(* Logix 5000 project; controller MV vendor 1 type 14 code 217 rev 31.11; software revision 31.00; part 35 of 53 *)
(* tags used below, declared in another part *)
   Alarm_Reset : BOOL;
   Analog_Fault_No : DINT;
   Analog_Simulation_Enabled : BOOL;
   CWD : CHECKWORD_FLAGS;
   Default_Check_Time : DINT;
   MV_MV18_RTD1_AI : PlantItem;   // MV18_RTD1
   MV_MV18_RTD1_AI_RawInput : ALIAS FOR Remote_IO:3:I.Ch5Data;   // Real Analog Input , Do Not Use In Code
   MV_MV19_RTD1_AI : PlantItem;   // MV19_RTD1
   MV_MV19_RTD1_AI_RawInput : ALIAS FOR Remote_IO:4:I.Ch0Data;   // Real Analog Input , Do Not Use In Code
   MV_MV20_RTD1_AI : PlantItem;   // MV20_RTD1
   MV_MV20_RTD1_AI_RawInput : ALIAS FOR Remote_IO:5:I.Ch1Data;   // Real Analog Input , Do Not Use In Code
   MV_MV21_RTD1_AI : PlantItem;   // MV21_RTD1
   MV_MV21_RTD1_AI_RawInput : ALIAS FOR Remote_IO:5:I.Ch2Data;   // Real Analog Input , Do Not Use In Code
   MV_MV22_RTD1_AI : PlantItem;   // MV22_RTD1
   MV_MV22_RTD1_AI_RawInput : ALIAS FOR Remote_IO:5:I.Ch3Data;   // Real Analog Input , Do Not Use In Code
   MV_MV23_RTD1_AI : PlantItem;   // MV23_RTD1
   MV_MV23_RTD1_AI_RawInput : ALIAS FOR Remote_IO:5:I.Ch4Data;   // Real Analog Input , Do Not Use In Code
   MV_MV30_RTD1_AI : PlantItem;   // MV30_RTD1
   MV_MV30_RTD1_AI_RawInput : ALIAS FOR Remote_IO:4:I.Ch1Data;   // Real Analog Input , Do Not Use In Code
   MV_MV31_RTD1_AI : PlantItem;   // MV31_RTD1
   MV_MV31_RTD1_AI_RawInput : ALIAS FOR Remote_IO:4:I.Ch2Data;   // Real Analog Input , Do Not Use In Code
   MV_MV32_RTD1_AI : PlantItem;   // MV32_RTD1
   MV_MV32_RTD1_AI_RawInput : ALIAS FOR Remote_IO:4:I.Ch3Data;   // Real Analog Input , Do Not Use In Code
   MV_MV33_RTD1_AI : PlantItem;   // MV33_RTD1
   MV_MV33_RTD1_AI_RawInput : ALIAS FOR Remote_IO:4:I.Ch4Data;   // Real Analog Input , Do Not Use In Code
   MV_MV34_RTD1_AI : PlantItem;   // MV34_RTD1
   MV_MV34_RTD1_AI_RawInput : ALIAS FOR Remote_IO:4:I.Ch5Data;   // Real Analog Input , Do Not Use In Code
   MV_MV35_RTD1_AI : PlantItem;   // MV35_RTD1
   MV_MV35_RTD1_AI_RawInput : ALIAS FOR Remote_IO:5:I.Ch0Data;   // Real Analog Input , Do Not Use In Code
   MV_MV36_TTX01_AI : PlantItem;   // MV36_TTX01
   MV_MV36_TTX01_AI_RawInput : ALIAS FOR Remote_IO:7:I.Ch00Data;   // Real Analog Input , Do Not Use In Code
   MV_MV37_TTX01_AI : PlantItem;   // MV37_TTX01
   MV_MV37_TTX01_AI_RawInput : ALIAS FOR Remote_IO:7:I.Ch01Data;   // Real Analog Input , Do Not Use In Code
   MV_MV38_TTX01_AI : PlantItem;   // MV38_TTX01
   MV_MV38_TTX01_AI_RawInput : ALIAS FOR Remote_IO:7:I.Ch02Data;   // Real Analog Input , Do Not Use In Code
   MV_MV39_TTX01_AI : PlantItem;   // MV39_TTX01
   MV_MV39_TTX01_AI_RawInput : ALIAS FOR Remote_IO:7:I.Ch03Data;   // Real Analog Input , Do Not Use In Code
   MV_MV40_TTX01_AI : PlantItem;   // MV40_TTX01
   MV_MV40_TTX01_AI_RawInput : ALIAS FOR Remote_IO:7:I.Ch04Data;   // Real Analog Input , Do Not Use In Code
   MV_MV41_TTX01_AI : PlantItem;   // MV41_TTX01
   MV_MV41_TTX01_AI_RawInput : ALIAS FOR Remote_IO:7:I.Ch05Data;   // Real Analog Input , Do Not Use In Code
   MV_MV42_TTX01_AI : PlantItem;   // MV42_TTX01
   MV_MV42_TTX01_AI_RawInput : ALIAS FOR Remote_IO:7:I.Ch06Data;   // Real Analog Input , Do Not Use In Code
   MV_MV43_TTX01_AI : PlantItem;   // MV43_TTX01
   MV_MV43_TTX01_AI_RawInput : ALIAS FOR Remote_IO:7:I.Ch07Data;   // Real Analog Input , Do Not Use In Code
   MV_MV44_TTX01_AI : PlantItem;   // MV44_TTX01
   MV_MV44_TTX01_AI_RawInput : ALIAS FOR Remote_IO:7:I.Ch08Data;   // Real Analog Input , Do Not Use In Code
   MV_MV45_TTX01_AI : PlantItem;   // MV45_TTX01
   MV_MV45_TTX01_AI_RawInput : ALIAS FOR Remote_IO:7:I.Ch09Data;   // Real Analog Input , Do Not Use In Code
   MV_MV46_TTX01_AI : PlantItem;   // MV46_TTX01
   MV_MV46_TTX01_AI_RawInput : ALIAS FOR Remote_IO:7:I.Ch10Data;   // Real Analog Input , Do Not Use In Code
   MV_MV47_TTX01_AI : PlantItem;   // MV47_TTX01
   MV_MV47_TTX01_AI_RawInput : ALIAS FOR Remote_IO:7:I.Ch11Data;   // Real Analog Input , Do Not Use In Code
   One_Second_One_Scan : ALIAS FOR One_Second_1_scan;
   overrange_RIO_analog_value : REAL;
   underrange_RIO_analog_value : REAL;
(* MV_Common, continued *)

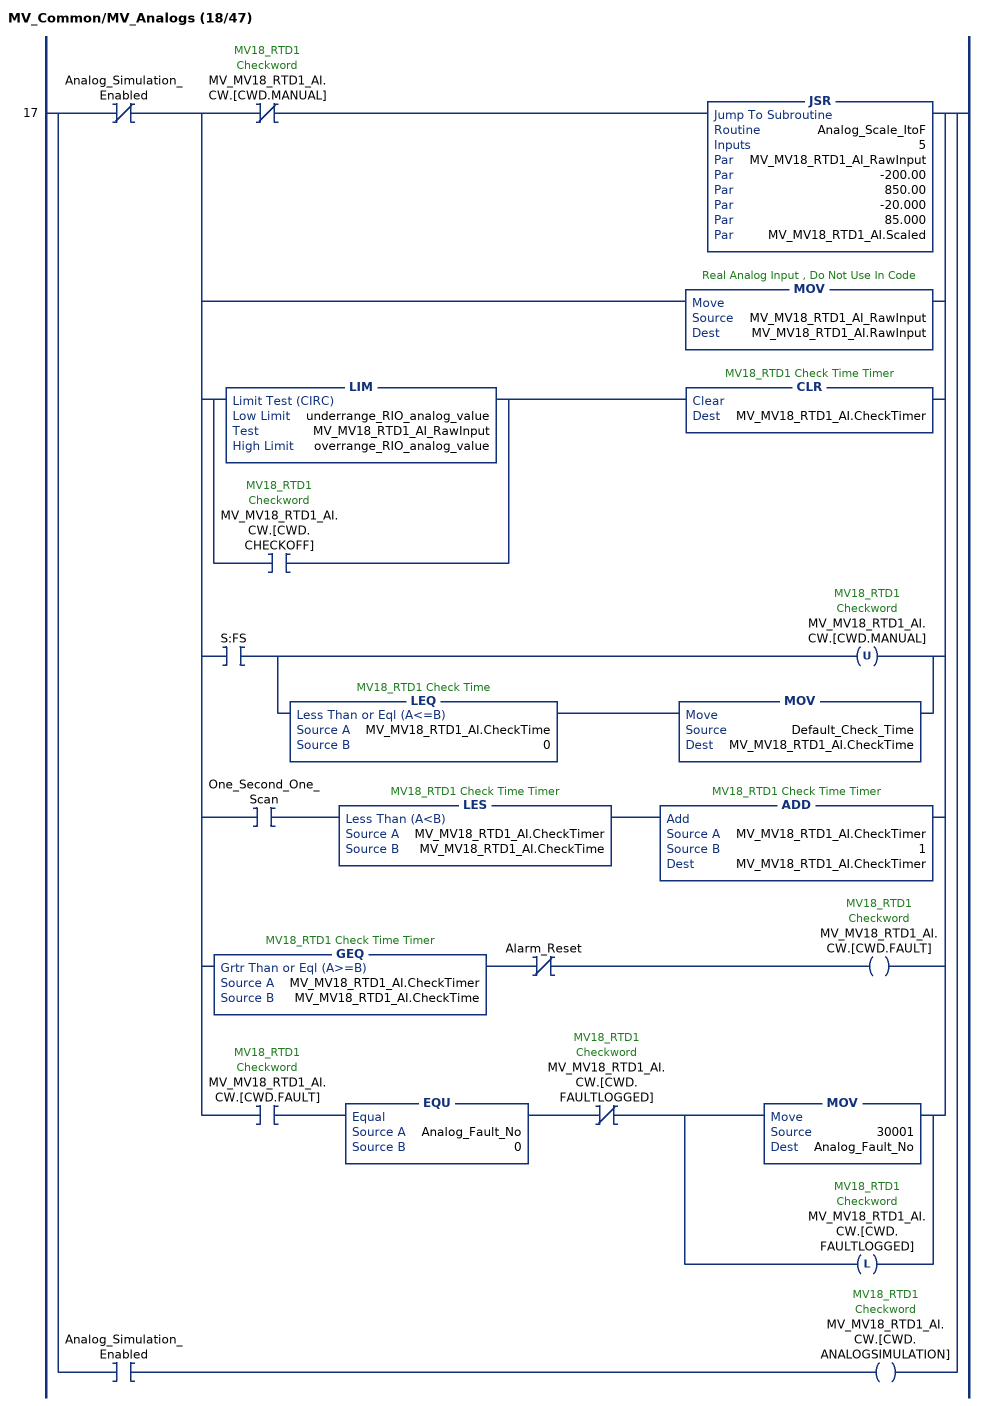
   [picture p810: MV_Common/MV_Analogs rungs 17-17]
   17: [XIO(Analog_Simulation_Enabled) [XIO(MV_MV18_RTD1_AI.CW.[CWD.MANUAL]) JSR(Analog_Scale_ItoF,5,MV_MV18_RTD1_AI_RawInput,-200.00,850.00,-20.000,85.000,MV_MV18_RTD1_AI.Scaled) ,MOV(MV_MV18_RTD1_AI_RawInput,MV_MV18_RTD1_AI.RawInput) ,[LIM(underrange_RIO_analog_value,MV_MV18_RTD1_AI_RawInput,overrange_RIO_analog_value) ,XIC(MV_MV18_RTD1_AI.CW.[CWD.CHECKOFF]) ] CLR(MV_MV18_RTD1_AI.CheckTimer) ,XIC(S:FS) [OTU(MV_MV18_RTD1_AI.CW.[CWD.MANUAL]) ,LEQ(MV_MV18_RTD1_AI.CheckTime,0) MOV(Default_Check_Time,MV_MV18_RTD1_AI.CheckTime) ] ,XIC(One_Second_One_Scan) LES(MV_MV18_RTD1_AI.CheckTimer,MV_MV18_RTD1_AI.CheckTime) ADD(MV_MV18_RTD1_AI.CheckTimer,1,MV_MV18_RTD1_AI.CheckTimer) ,GEQ(MV_MV18_RTD1_AI.CheckTimer,MV_MV18_RTD1_AI.CheckTime) XIO(Alarm_Reset) OTE(MV_MV18_RTD1_AI.CW.[CWD.FAULT]) ,XIC(MV_MV18_RTD1_AI.CW.[CWD.FAULT]) EQU(Analog_Fault_No,0) XIO(MV_MV18_RTD1_AI.CW.[CWD.FAULTLOGGED]) [MOV(30001,Analog_Fault_No) ,OTL(MV_MV18_RTD1_AI.CW.[CWD.FAULTLOGGED]) ] ] ,XIC(Analog_Simulation_Enabled) OTE(MV_MV18_RTD1_AI.CW.[CWD.ANALOGSIMULATION]) ];
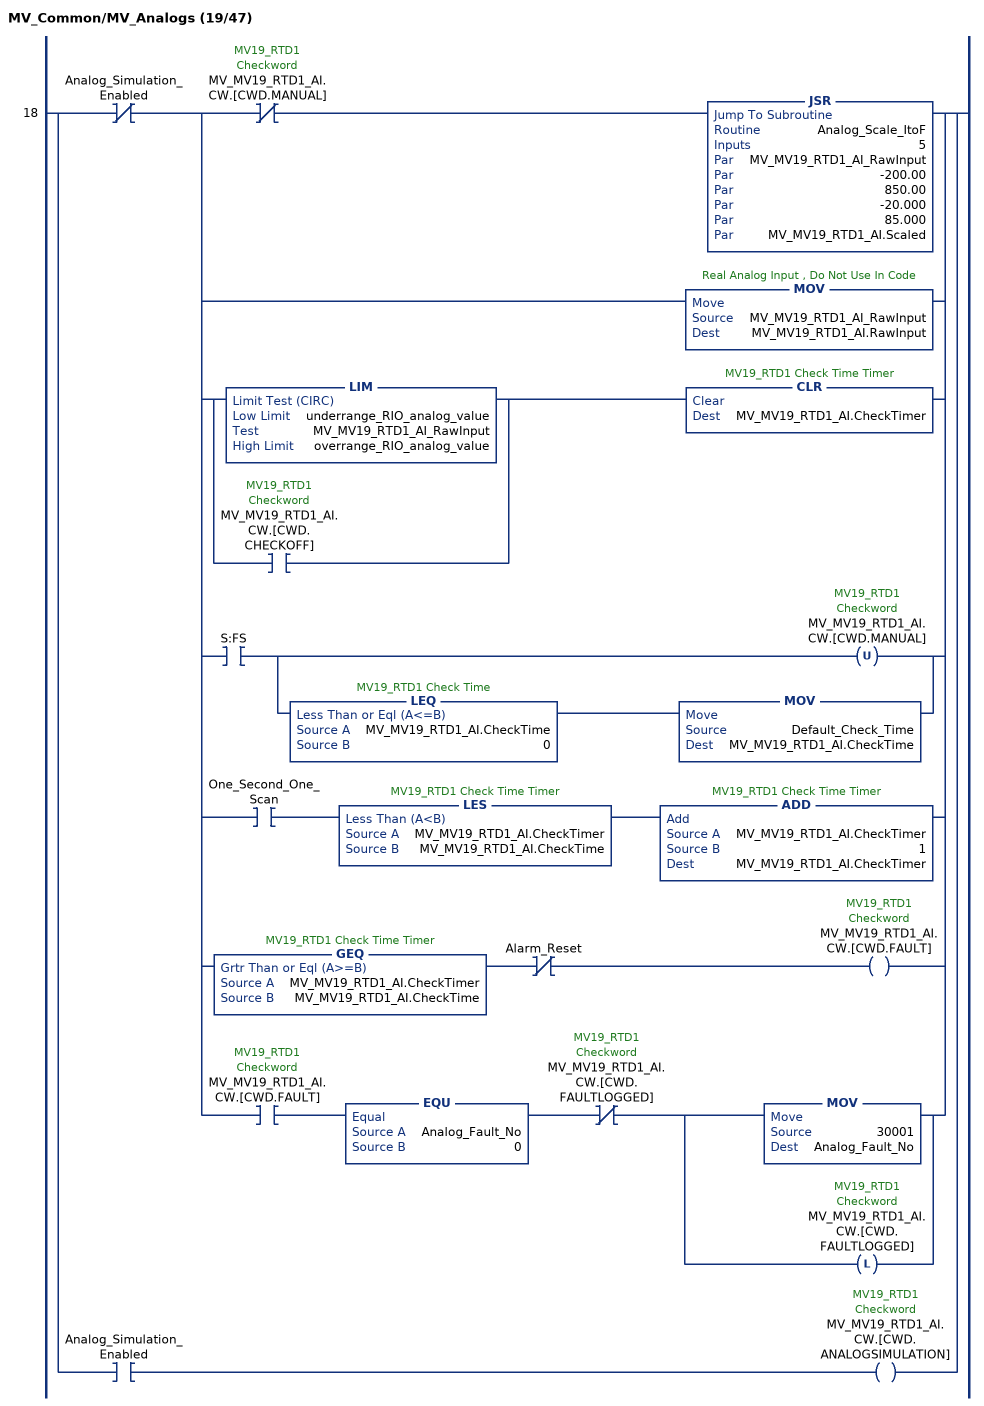
   18: [XIO(Analog_Simulation_Enabled) [XIO(MV_MV19_RTD1_AI.CW.[CWD.MANUAL]) JSR(Analog_Scale_ItoF,5,MV_MV19_RTD1_AI_RawInput,-200.00,850.00,-20.000,85.000,MV_MV19_RTD1_AI.Scaled) ,MOV(MV_MV19_RTD1_AI_RawInput,MV_MV19_RTD1_AI.RawInput) ,[LIM(underrange_RIO_analog_value,MV_MV19_RTD1_AI_RawInput,overrange_RIO_analog_value) ,XIC(MV_MV19_RTD1_AI.CW.[CWD.CHECKOFF]) ] CLR(MV_MV19_RTD1_AI.CheckTimer) ,XIC(S:FS) [OTU(MV_MV19_RTD1_AI.CW.[CWD.MANUAL]) ,LEQ(MV_MV19_RTD1_AI.CheckTime,0) MOV(Default_Check_Time,MV_MV19_RTD1_AI.CheckTime) ] ,XIC(One_Second_One_Scan) LES(MV_MV19_RTD1_AI.CheckTimer,MV_MV19_RTD1_AI.CheckTime) ADD(MV_MV19_RTD1_AI.CheckTimer,1,MV_MV19_RTD1_AI.CheckTimer) ,GEQ(MV_MV19_RTD1_AI.CheckTimer,MV_MV19_RTD1_AI.CheckTime) XIO(Alarm_Reset) OTE(MV_MV19_RTD1_AI.CW.[CWD.FAULT]) ,XIC(MV_MV19_RTD1_AI.CW.[CWD.FAULT]) EQU(Analog_Fault_No,0) XIO(MV_MV19_RTD1_AI.CW.[CWD.FAULTLOGGED]) [MOV(30001,Analog_Fault_No) ,OTL(MV_MV19_RTD1_AI.CW.[CWD.FAULTLOGGED]) ] ] ,XIC(Analog_Simulation_Enabled) OTE(MV_MV19_RTD1_AI.CW.[CWD.ANALOGSIMULATION]) ];
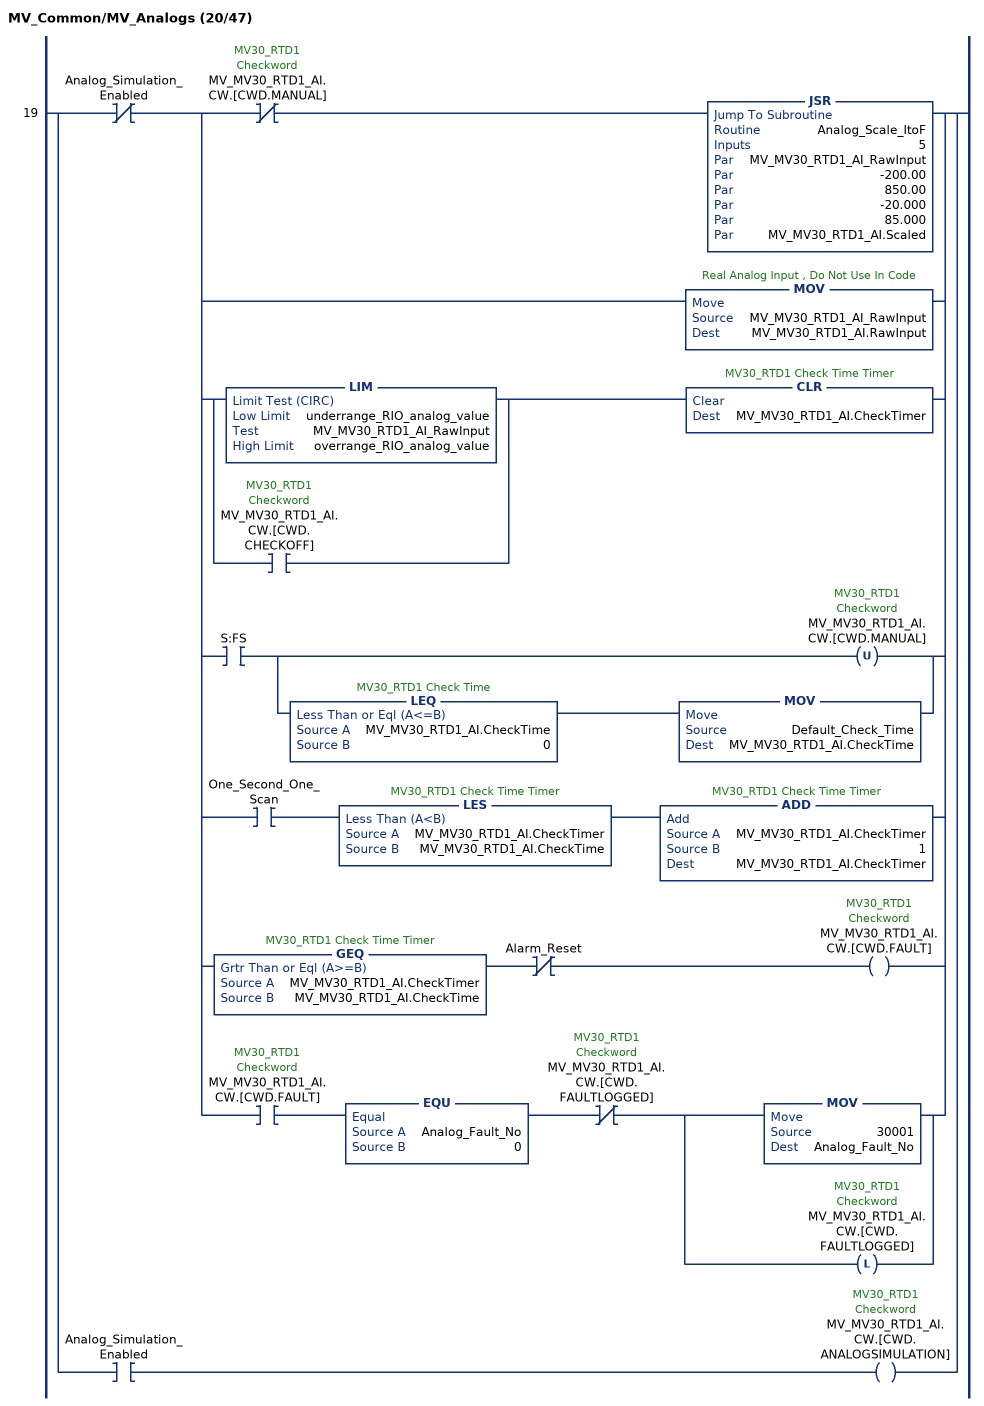
   19: [XIO(Analog_Simulation_Enabled) [XIO(MV_MV30_RTD1_AI.CW.[CWD.MANUAL]) JSR(Analog_Scale_ItoF,5,MV_MV30_RTD1_AI_RawInput,-200.00,850.00,-20.000,85.000,MV_MV30_RTD1_AI.Scaled) ,MOV(MV_MV30_RTD1_AI_RawInput,MV_MV30_RTD1_AI.RawInput) ,[LIM(underrange_RIO_analog_value,MV_MV30_RTD1_AI_RawInput,overrange_RIO_analog_value) ,XIC(MV_MV30_RTD1_AI.CW.[CWD.CHECKOFF]) ] CLR(MV_MV30_RTD1_AI.CheckTimer) ,XIC(S:FS) [OTU(MV_MV30_RTD1_AI.CW.[CWD.MANUAL]) ,LEQ(MV_MV30_RTD1_AI.CheckTime,0) MOV(Default_Check_Time,MV_MV30_RTD1_AI.CheckTime) ] ,XIC(One_Second_One_Scan) LES(MV_MV30_RTD1_AI.CheckTimer,MV_MV30_RTD1_AI.CheckTime) ADD(MV_MV30_RTD1_AI.CheckTimer,1,MV_MV30_RTD1_AI.CheckTimer) ,GEQ(MV_MV30_RTD1_AI.CheckTimer,MV_MV30_RTD1_AI.CheckTime) XIO(Alarm_Reset) OTE(MV_MV30_RTD1_AI.CW.[CWD.FAULT]) ,XIC(MV_MV30_RTD1_AI.CW.[CWD.FAULT]) EQU(Analog_Fault_No,0) XIO(MV_MV30_RTD1_AI.CW.[CWD.FAULTLOGGED]) [MOV(30001,Analog_Fault_No) ,OTL(MV_MV30_RTD1_AI.CW.[CWD.FAULTLOGGED]) ] ] ,XIC(Analog_Simulation_Enabled) OTE(MV_MV30_RTD1_AI.CW.[CWD.ANALOGSIMULATION]) ];
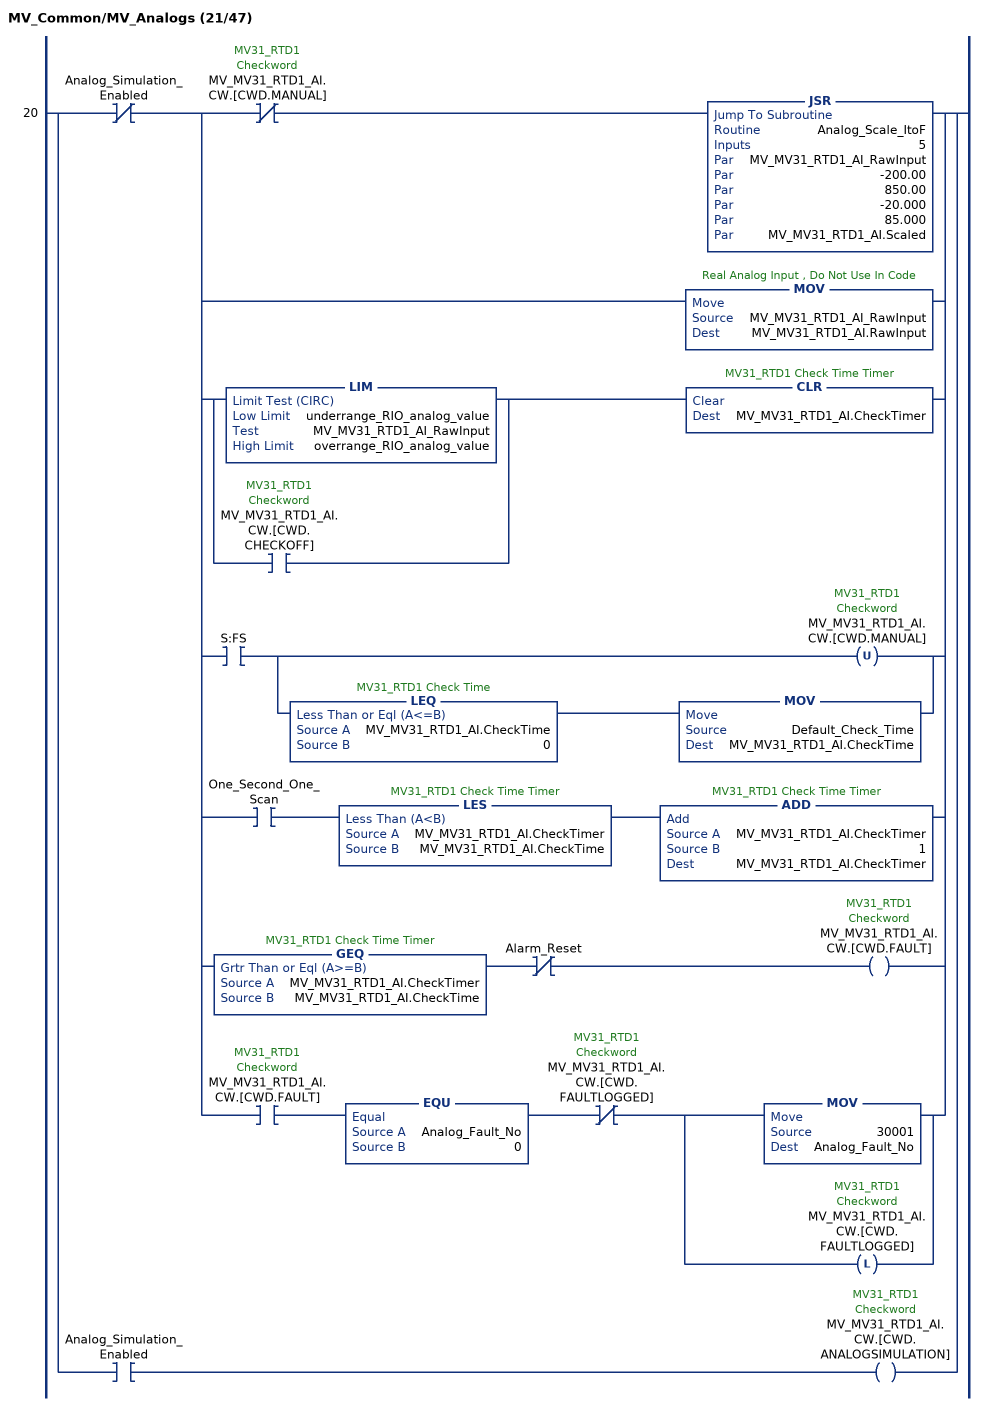
   20: [XIO(Analog_Simulation_Enabled) [XIO(MV_MV31_RTD1_AI.CW.[CWD.MANUAL]) JSR(Analog_Scale_ItoF,5,MV_MV31_RTD1_AI_RawInput,-200.00,850.00,-20.000,85.000,MV_MV31_RTD1_AI.Scaled) ,MOV(MV_MV31_RTD1_AI_RawInput,MV_MV31_RTD1_AI.RawInput) ,[LIM(underrange_RIO_analog_value,MV_MV31_RTD1_AI_RawInput,overrange_RIO_analog_value) ,XIC(MV_MV31_RTD1_AI.CW.[CWD.CHECKOFF]) ] CLR(MV_MV31_RTD1_AI.CheckTimer) ,XIC(S:FS) [OTU(MV_MV31_RTD1_AI.CW.[CWD.MANUAL]) ,LEQ(MV_MV31_RTD1_AI.CheckTime,0) MOV(Default_Check_Time,MV_MV31_RTD1_AI.CheckTime) ] ,XIC(One_Second_One_Scan) LES(MV_MV31_RTD1_AI.CheckTimer,MV_MV31_RTD1_AI.CheckTime) ADD(MV_MV31_RTD1_AI.CheckTimer,1,MV_MV31_RTD1_AI.CheckTimer) ,GEQ(MV_MV31_RTD1_AI.CheckTimer,MV_MV31_RTD1_AI.CheckTime) XIO(Alarm_Reset) OTE(MV_MV31_RTD1_AI.CW.[CWD.FAULT]) ,XIC(MV_MV31_RTD1_AI.CW.[CWD.FAULT]) EQU(Analog_Fault_No,0) XIO(MV_MV31_RTD1_AI.CW.[CWD.FAULTLOGGED]) [MOV(30001,Analog_Fault_No) ,OTL(MV_MV31_RTD1_AI.CW.[CWD.FAULTLOGGED]) ] ] ,XIC(Analog_Simulation_Enabled) OTE(MV_MV31_RTD1_AI.CW.[CWD.ANALOGSIMULATION]) ];
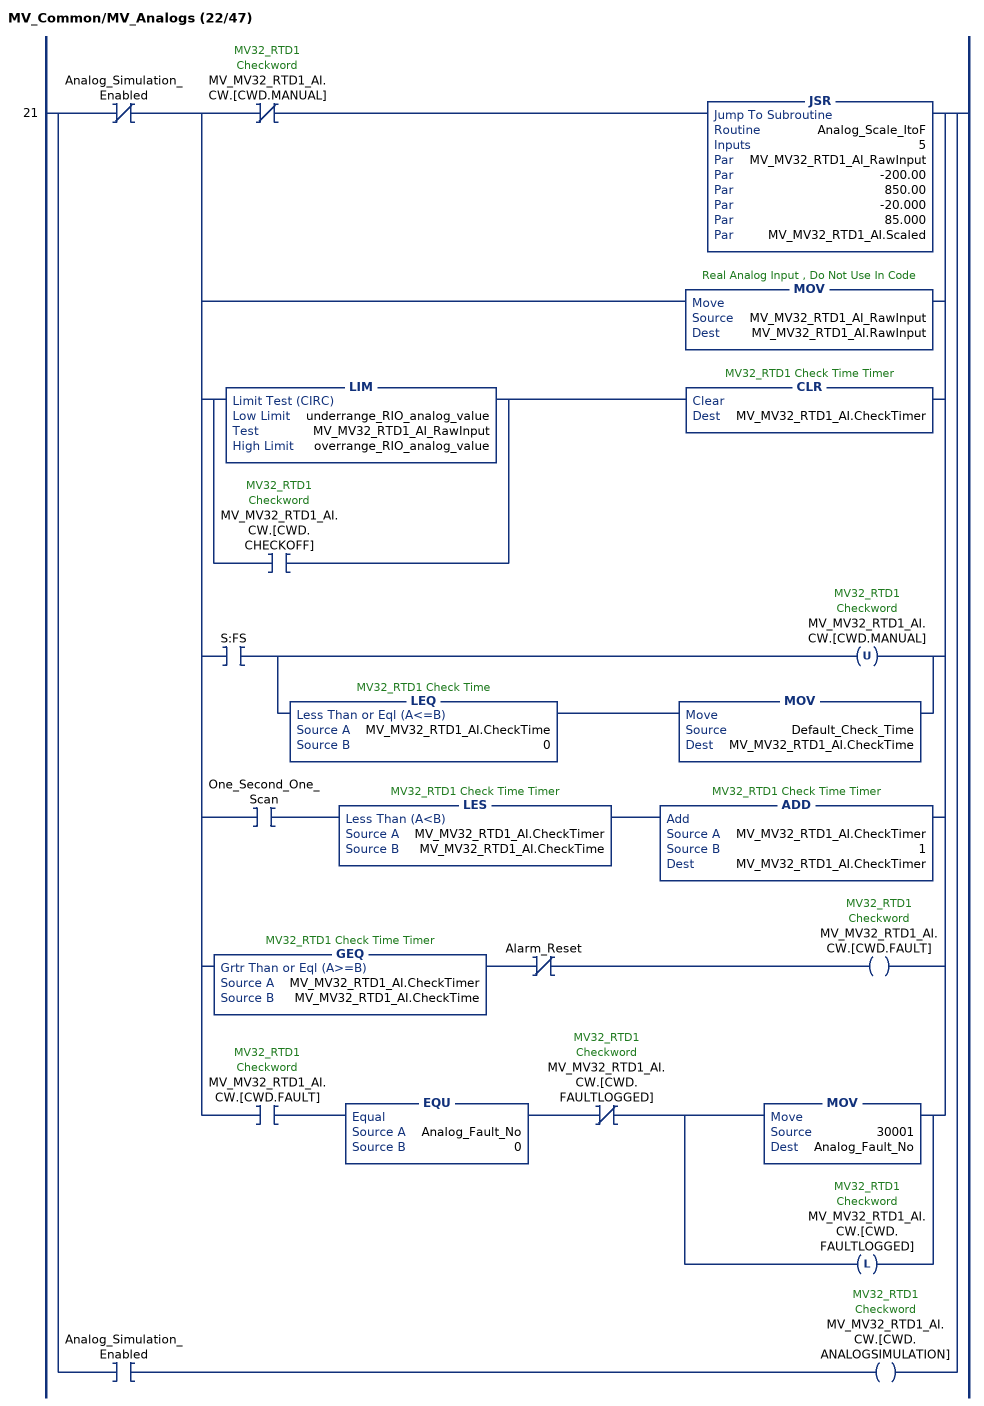
   21: [XIO(Analog_Simulation_Enabled) [XIO(MV_MV32_RTD1_AI.CW.[CWD.MANUAL]) JSR(Analog_Scale_ItoF,5,MV_MV32_RTD1_AI_RawInput,-200.00,850.00,-20.000,85.000,MV_MV32_RTD1_AI.Scaled) ,MOV(MV_MV32_RTD1_AI_RawInput,MV_MV32_RTD1_AI.RawInput) ,[LIM(underrange_RIO_analog_value,MV_MV32_RTD1_AI_RawInput,overrange_RIO_analog_value) ,XIC(MV_MV32_RTD1_AI.CW.[CWD.CHECKOFF]) ] CLR(MV_MV32_RTD1_AI.CheckTimer) ,XIC(S:FS) [OTU(MV_MV32_RTD1_AI.CW.[CWD.MANUAL]) ,LEQ(MV_MV32_RTD1_AI.CheckTime,0) MOV(Default_Check_Time,MV_MV32_RTD1_AI.CheckTime) ] ,XIC(One_Second_One_Scan) LES(MV_MV32_RTD1_AI.CheckTimer,MV_MV32_RTD1_AI.CheckTime) ADD(MV_MV32_RTD1_AI.CheckTimer,1,MV_MV32_RTD1_AI.CheckTimer) ,GEQ(MV_MV32_RTD1_AI.CheckTimer,MV_MV32_RTD1_AI.CheckTime) XIO(Alarm_Reset) OTE(MV_MV32_RTD1_AI.CW.[CWD.FAULT]) ,XIC(MV_MV32_RTD1_AI.CW.[CWD.FAULT]) EQU(Analog_Fault_No,0) XIO(MV_MV32_RTD1_AI.CW.[CWD.FAULTLOGGED]) [MOV(30001,Analog_Fault_No) ,OTL(MV_MV32_RTD1_AI.CW.[CWD.FAULTLOGGED]) ] ] ,XIC(Analog_Simulation_Enabled) OTE(MV_MV32_RTD1_AI.CW.[CWD.ANALOGSIMULATION]) ];
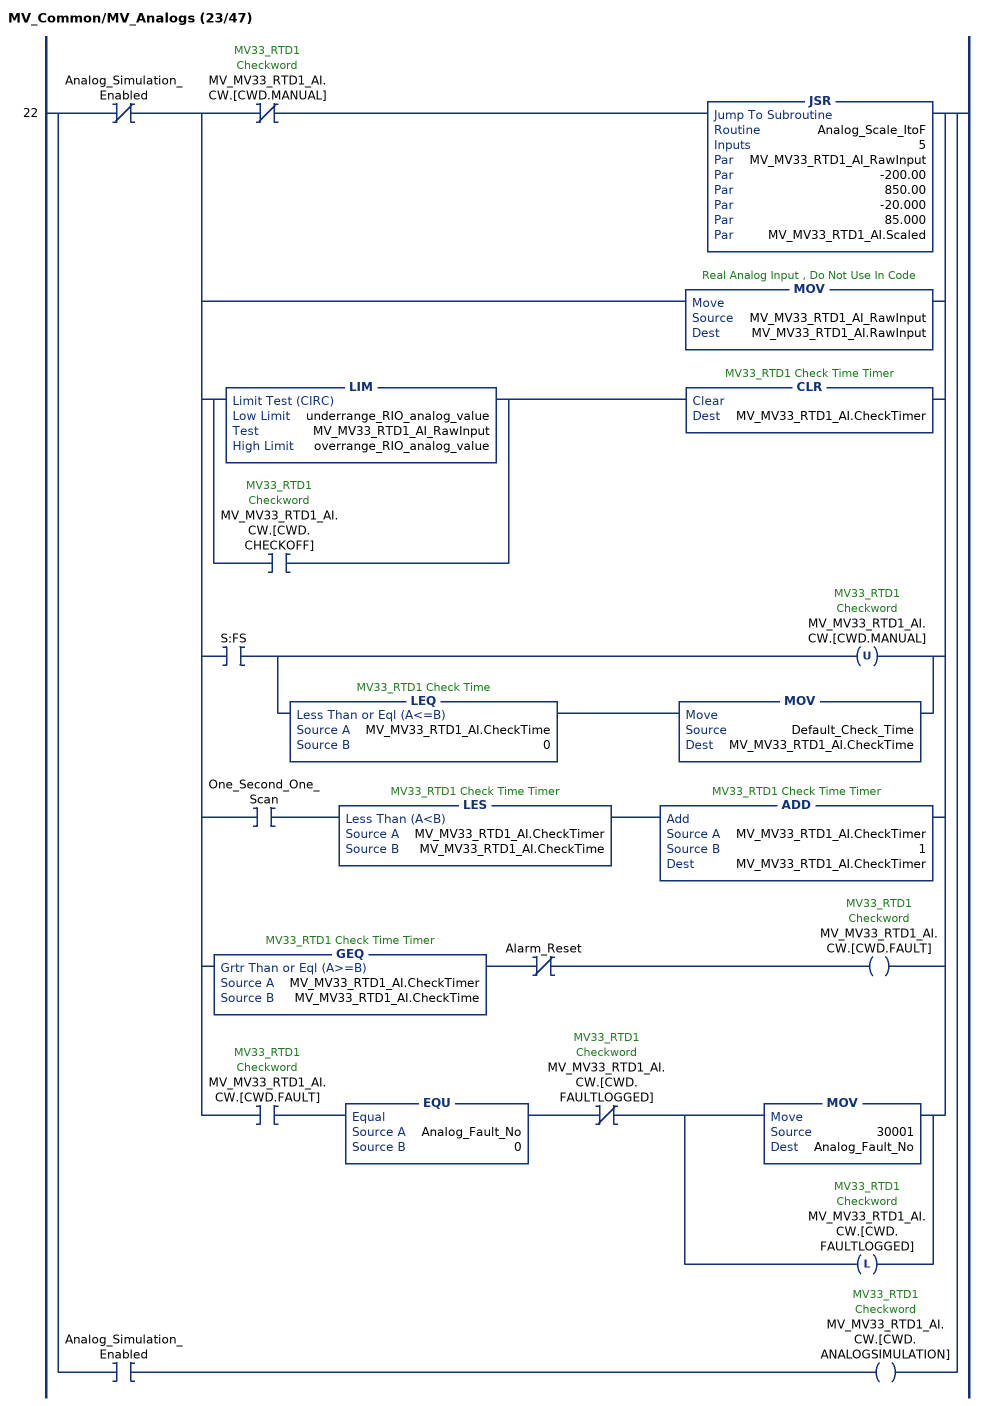
   22: [XIO(Analog_Simulation_Enabled) [XIO(MV_MV33_RTD1_AI.CW.[CWD.MANUAL]) JSR(Analog_Scale_ItoF,5,MV_MV33_RTD1_AI_RawInput,-200.00,850.00,-20.000,85.000,MV_MV33_RTD1_AI.Scaled) ,MOV(MV_MV33_RTD1_AI_RawInput,MV_MV33_RTD1_AI.RawInput) ,[LIM(underrange_RIO_analog_value,MV_MV33_RTD1_AI_RawInput,overrange_RIO_analog_value) ,XIC(MV_MV33_RTD1_AI.CW.[CWD.CHECKOFF]) ] CLR(MV_MV33_RTD1_AI.CheckTimer) ,XIC(S:FS) [OTU(MV_MV33_RTD1_AI.CW.[CWD.MANUAL]) ,LEQ(MV_MV33_RTD1_AI.CheckTime,0) MOV(Default_Check_Time,MV_MV33_RTD1_AI.CheckTime) ] ,XIC(One_Second_One_Scan) LES(MV_MV33_RTD1_AI.CheckTimer,MV_MV33_RTD1_AI.CheckTime) ADD(MV_MV33_RTD1_AI.CheckTimer,1,MV_MV33_RTD1_AI.CheckTimer) ,GEQ(MV_MV33_RTD1_AI.CheckTimer,MV_MV33_RTD1_AI.CheckTime) XIO(Alarm_Reset) OTE(MV_MV33_RTD1_AI.CW.[CWD.FAULT]) ,XIC(MV_MV33_RTD1_AI.CW.[CWD.FAULT]) EQU(Analog_Fault_No,0) XIO(MV_MV33_RTD1_AI.CW.[CWD.FAULTLOGGED]) [MOV(30001,Analog_Fault_No) ,OTL(MV_MV33_RTD1_AI.CW.[CWD.FAULTLOGGED]) ] ] ,XIC(Analog_Simulation_Enabled) OTE(MV_MV33_RTD1_AI.CW.[CWD.ANALOGSIMULATION]) ];
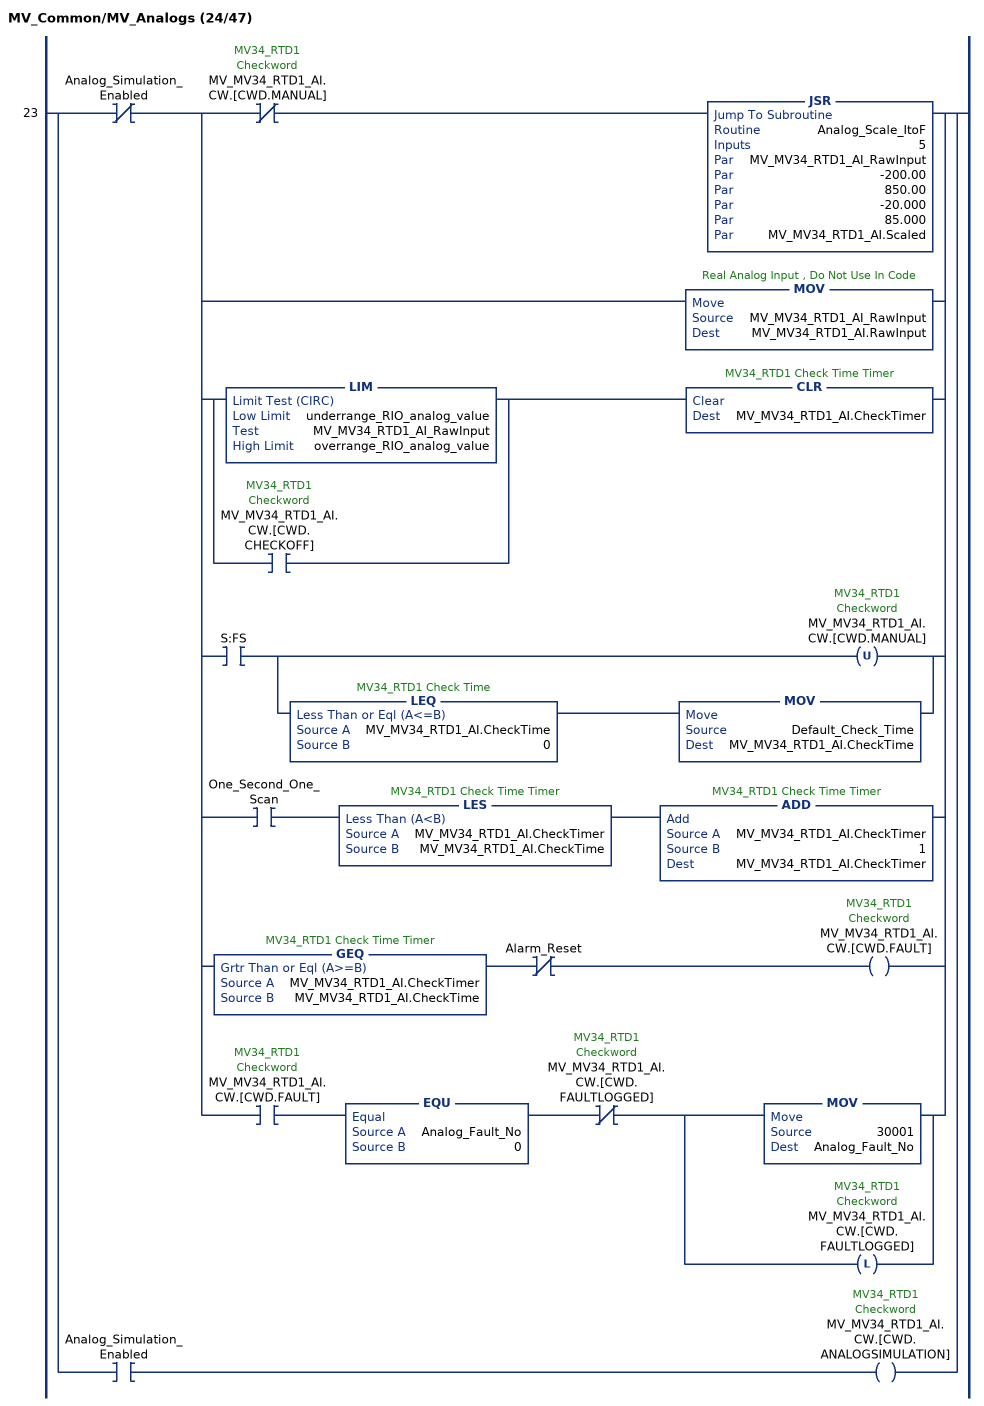
   23: [XIO(Analog_Simulation_Enabled) [XIO(MV_MV34_RTD1_AI.CW.[CWD.MANUAL]) JSR(Analog_Scale_ItoF,5,MV_MV34_RTD1_AI_RawInput,-200.00,850.00,-20.000,85.000,MV_MV34_RTD1_AI.Scaled) ,MOV(MV_MV34_RTD1_AI_RawInput,MV_MV34_RTD1_AI.RawInput) ,[LIM(underrange_RIO_analog_value,MV_MV34_RTD1_AI_RawInput,overrange_RIO_analog_value) ,XIC(MV_MV34_RTD1_AI.CW.[CWD.CHECKOFF]) ] CLR(MV_MV34_RTD1_AI.CheckTimer) ,XIC(S:FS) [OTU(MV_MV34_RTD1_AI.CW.[CWD.MANUAL]) ,LEQ(MV_MV34_RTD1_AI.CheckTime,0) MOV(Default_Check_Time,MV_MV34_RTD1_AI.CheckTime) ] ,XIC(One_Second_One_Scan) LES(MV_MV34_RTD1_AI.CheckTimer,MV_MV34_RTD1_AI.CheckTime) ADD(MV_MV34_RTD1_AI.CheckTimer,1,MV_MV34_RTD1_AI.CheckTimer) ,GEQ(MV_MV34_RTD1_AI.CheckTimer,MV_MV34_RTD1_AI.CheckTime) XIO(Alarm_Reset) OTE(MV_MV34_RTD1_AI.CW.[CWD.FAULT]) ,XIC(MV_MV34_RTD1_AI.CW.[CWD.FAULT]) EQU(Analog_Fault_No,0) XIO(MV_MV34_RTD1_AI.CW.[CWD.FAULTLOGGED]) [MOV(30001,Analog_Fault_No) ,OTL(MV_MV34_RTD1_AI.CW.[CWD.FAULTLOGGED]) ] ] ,XIC(Analog_Simulation_Enabled) OTE(MV_MV34_RTD1_AI.CW.[CWD.ANALOGSIMULATION]) ];